FUNCTION_BLOCK "FB_BreakDetector_V1.00"   // FB20, LAD
{ S7_Optimized_Access := 'TRUE' }
VERSION : 0.1
   VAR_INPUT
      IN_xCycleON : Bool;   // Cycle ON
      IN_xCycleONDel : Bool;   // Delayed cycle ON signal
      IN_xGeneralReset : Bool;   // General reset
      IN_xResetAlarms : Bool;   // Reset alarms
      IN_xFaultsEnabled : Bool;   // Faults enabled
      IN_dNumUsedPhoto : DInt;   // Number of used photocell
      IN_dIndexBreakMachine : DInt;   // Index break machine on buffer
      INPUT : Struct   // Digital inputs
         xPowerSupplyControl : Bool;   // Power supply control
         xConnectorONOp : Bool;   // Control connector ON operator side
         xConnectorONOppoOp : Bool;   // Control connector ON opposite operator side
         xButtonAlarmOFF : Bool;   // Reset horn alarm
         rgxPhotoStatus : Array[0..#CONST_DMAXPHOTOCELL_IND] of Bool;   // Photocell status
      END_STRUCT;
   END_VAR
   VAR_OUTPUT
      OUTPUT : Struct
         xLampBreakAlarm : Bool;   // HL.Break alam
         xSirenBreakAlarm : Bool;   // HA.Break alam
      END_STRUCT;
   END_VAR
   VAR_IN_OUT
      INO_tEncoder : "UDT_Encoder";   // Encoder data
      INO_tRibbon : "UDT_RibbonData";   // Ribbona data
      INO_tFBAddDefect : "FB_Defects_Add_V1.00";   // Add defect
      INO_xDefectBufferFull : Bool;   // Defect buffer full
   END_VAR
   VAR RETAIN
      tHMW : Struct   // HMI Write
         dMinBreakSize_cmm : DInt;   // Minimum breaksize [mm/100] {mm/100|mm|0|1000|O}
         rgxEnabledPhotocell : Array[0..#CONST_DMAXPHOTOCELL_IND] of Bool;   // Photocell abilitation (1=Disabled 3=Enabled) {X|X|X|X|O}
         dDistanceSnaproll_cmm : DInt;   // Distance from snaproll [mm/100] {mm/100|mm|0|60000|O}
         xUpdateDistanceSnap : Bool;   // Update distance from snaproll {X|X|X|X|O}
      END_STRUCT;
      tHMR : Struct   // HMI Read
         dStatus : DInt;   // Status (1=Idle 3=Run 5= Glass break 7=Anomaly) {X|X|X|X|O}
         dDistanceSnaproll_cmm : DInt;   // Distance from snaproll [mm/100] {mm/100|mm|0|60000|O}
         rgxPhotoStatus : Array[0..#CONST_DMAXPHOTOCELL_IND] of Bool;   // Photocell status (0=OFF 1=ON) {X|X|X|X|O}
         rgdPhotoAbilitation : Array[0..#CONST_DMAXPHOTOCELL_IND] of DInt;   // Photocell abilitation (1=Disabled 3=Enabled) {X|X|X|X|O}
      END_STRUCT;
   END_VAR
   VAR
      tALM : Struct   // HMI Alarms
         tS : Struct   // Stopping faults machine
            xPowerSupplyControl : Bool;   // Power supply control {X|X|X|X|O}
            xConnectorONOpSide : Bool;   // Connector ON operator side {X|X|X|X|O}
            xConnectorONOppoOpSide : Bool;   // Connector ON opposite operator side {X|X|X|X|O}
            xSpare_3 : Bool;
            xSpare_4 : Bool;
            xSpare_5 : Bool;
            xSpare_6 : Bool;
            xSpare_7 : Bool;
            xSpare_8 : Bool;
            xSpare_9 : Bool;
            xSpare_10 : Bool;
            xSpare_11 : Bool;
            xSpare_12 : Bool;
            xSpare_13 : Bool;
            xSpare_14 : Bool;
            xSpare_15 : Bool;
            xSpare_16 : Bool;
            xSpare_17 : Bool;
            xSpare_18 : Bool;
            xSpare_19 : Bool;
            xSpare_20 : Bool;
            xSpare_21 : Bool;
            xSpare_22 : Bool;
            xSpare_23 : Bool;
            xSpare_24 : Bool;
            xSpare_25 : Bool;
            xSpare_26 : Bool;
            xSpare_27 : Bool;
            xSpare_28 : Bool;
            xSpare_29 : Bool;
            xSpare_30 : Bool;
            xSpare_31 : Bool;
         END_STRUCT;
         tF : Struct   // Faults
            xGlassBreakPhotocell1 : Bool;   // Glass break on photocell #1
            xGlassBreakPhotocell2 : Bool;   // Glass break on photocell #2
            xGlassBreakPhotocell3 : Bool;   // Glass break on photocell #3
            xGlassBreakPhotocell4 : Bool;   // Glass break on photocell #4
            xGlassBreakPhotocell5 : Bool;   // Glass break on photocell #5
            xGlassBreakPhotocell6 : Bool;   // Glass break on photocell #6
            xGlassBreakPhotocell7 : Bool;   // Glass break on photocell #7
            xGlassBreakPhotocell8 : Bool;   // Glass break on photocell #8
            xGlassBreakPhotocell9 : Bool;   // Glass break on photocell #9
            xGlassBreakPhotocell10 : Bool;   // Glass break on photocell #10
            xGlassBreakPhotocell11 : Bool;   // Glass break on photocell #11
            xGlassBreakPhotocell12 : Bool;   // Glass break on photocell #12
            xGlassBreakPhotocell13 : Bool;   // Glass break on photocell #13
            xGlassBreakPhotocell14 : Bool;   // Glass break on photocell #14
            xGlassBreakPhotocell15 : Bool;   // Glass break on photocell #15
            xGlassBreakPhotocell16 : Bool;   // Glass break on photocell #16
            xGlassBreakPhotocell17 : Bool;   // Glass break on photocell #17
            xGlassBreakPhotocell18 : Bool;   // Glass break on photocell #18
            xGlassBreakPhotocell19 : Bool;   // Glass break on photocell #19
            xGlassBreakPhotocell20 : Bool;   // Glass break on photocell #20
            xGlassBreakPhotocell21 : Bool;   // Glass break on photocell #21
            xGlassBreakPhotocell22 : Bool;   // Glass break on photocell #22
            xGlassBreakPhotocell23 : Bool;   // Glass break on photocell #23
            xGlassBreakPhotocell24 : Bool;   // Glass break on photocell #24
            xGlassBreakPhotocell25 : Bool;   // Glass break on photocell #25
            xGlassBreakPhotocell26 : Bool;   // Glass break on photocell #26
            xGlassBreakPhotocell27 : Bool;   // Glass break on photocell #27
            xGlassBreakPhotocell28 : Bool;   // Glass break on photocell #28
            xGlassBreakPhotocell29 : Bool;   // Glass break on photocell #29
            xGlassBreakPhotocell30 : Bool;   // Glass break on photocell #30
            xGlassBreakPhotocell31 : Bool;   // Glass break on photocell #31
            xGlassBreakPhotocell32 : Bool;   // Glass break on photocell #32
         END_STRUCT;
         tW : Struct   // Warnings
            xSpare_0 : Bool;
            xSpare_1 : Bool;
            xSpare_2 : Bool;
            xSpare_3 : Bool;
            xSpare_4 : Bool;
            xSpare_5 : Bool;
            xSpare_6 : Bool;
            xSpare_7 : Bool;
            xSpare_8 : Bool;
            xSpare_9 : Bool;
            xSpare_10 : Bool;
            xSpare_11 : Bool;
            xSpare_12 : Bool;
            xSpare_13 : Bool;
            xSpare_14 : Bool;
            xSpare_15 : Bool;
            xSpare_16 : Bool;
            xSpare_17 : Bool;
            xSpare_18 : Bool;
            xSpare_19 : Bool;
            xSpare_20 : Bool;
            xSpare_21 : Bool;
            xSpare_22 : Bool;
            xSpare_23 : Bool;
            xSpare_24 : Bool;
            xSpare_25 : Bool;
            xSpare_26 : Bool;
            xSpare_27 : Bool;
            xSpare_28 : Bool;
            xSpare_29 : Bool;
            xSpare_30 : Bool;
            xSpare_31 : Bool;
         END_STRUCT;
      END_STRUCT;
      ST_xOutputEnable : Bool;   // Output enable
      ST_xStoppedFaults : Bool;   // Stopped faults
      ST_xFaults : Bool;   // Faults
      ST_xWarning : Bool;   // Warnings
      AUX_rgxLastPhotoState : Array[0..#CONST_DMAXPHOTOCELL_IND] of Bool;   // Last photocell status
      AUX_xGlassBreak : Bool;   // Glass break in progress
      AUX_xGlassBreakInGoing : Bool;   // Glass break ingoing
      AUX_dCounterOnBreak_cmm : DInt;   // Encoder counter on glass break front
      AUX_dLastInsertDefectPos_cmm : DInt;   // Last inserted defect position [mm/100]
      OSR_xGlassBreak : Bool;   // OSR glasss break
   END_VAR
   VAR_TEMP
      TMP_dwValue : DWord;
      TMP_dIndex : DInt;
      TMP_dNumUsedPhotocell : DInt;
      TMP_xGlassBreak : Bool;
      TMP_xAtLeastOnePhoto : Bool;
      TMP_dEncDef_cmm : DInt;
   END_VAR
   VAR CONSTANT
      CONST_DMAXPHOTOCELL : DInt := 32;   // Maximum number of photocell
      CONST_DMAXPHOTOCELL_IND : DInt := 31;   // Maximum number of photocell index (Always -1)
      CONST_DGLASSBREAK_CLASS : DInt := 21;   // Glass break used class
      CONST_DGLASSBREAK_SUBTYPE : DInt := 1002;   // Glass break subtype
      CONST_DGLASSBREAK_DEFECT_WIDTH_CMM : DInt := 366000;   // Defect width [mm/100]
      CONST_DGLASSBREAK_DEFECT_GAP_CMM : DInt := 40000;   // Glass break defect gap [mm/100]
      CONST_DGLASSBREAK_LASTDEFECT_LENGTH_CMM : DInt := 50000;   // Last defect on glass break length [mm/100]
   END_VAR
   VAR_TEMP   // added for the SCL form of the ladder/FBD networks
      _w1 : Bool;
   END_VAR
BEGIN

REGION Network 1: ####_CONSTANTS_####
END_REGION

REGION Network 2: ####_MATCH_####
END_REGION

REGION Network 3 (SCL): ### SIMULATION ###
   IF "SIMULATION_ACTIVE" THEN
       #INPUT.xConnectorONOp := TRUE;
       #INPUT.xConnectorONOppoOp := TRUE;
       #INPUT.xPowerSupplyControl := TRUE;
    //   #INPUT.rgxPhotoStatus[0] := 1;
   //    #INPUT.rgxPhotoStatus[1] := 1;
   //    #INPUT.rgxPhotoStatus[2] := 1;
   //    #INPUT.rgxPhotoStatus[3] := 1;
    //   #INPUT.rgxPhotoStatus[4] := 1;
     //  #INPUT.rgxPhotoStatus[5] := 1;
    //   #INPUT.rgxPhotoStatus[6] := 1;
     //  #INPUT.rgxPhotoStatus[7] := 1;
     //  #INPUT.rgxPhotoStatus[8] := 1;
      // #INPUT.rgxPhotoStatus[9] := 1;
   END_IF;
END_REGION

REGION Network 4 (SCL): Evaluate number of used photocell
   #TMP_dNumUsedPhotocell := #IN_dNumUsedPhoto;

   IF #TMP_dNumUsedPhotocell > #CONST_DMAXPHOTOCELL THEN
       #TMP_dNumUsedPhotocell := #CONST_DMAXPHOTOCELL;
   ELSIF #TMP_dNumUsedPhotocell < 0 THEN
       #TMP_dNumUsedPhotocell := 0;
   END_IF;
END_REGION

REGION Network 5 (SCL): Reset all the pending status
   IF #IN_xGeneralReset THEN
       #AUX_xGlassBreak := FALSE;
       #AUX_xGlassBreakInGoing := FALSE;
       #AUX_dCounterOnBreak_cmm := 0;

       FOR #TMP_dIndex := 0 TO #TMP_dNumUsedPhotocell - 1 DO
           #AUX_rgxLastPhotoState[#TMP_dIndex] := FALSE;
       END_FOR;

   END_IF;
END_REGION

REGION Network 6: ####_HMI_LOGICS_####
END_REGION

REGION Network 7 (SCL): Manage HMI Logics
   FOR #TMP_dIndex := 0 TO #TMP_dNumUsedPhotocell - 1 DO

       (*  IF #tHMW.rgxEnabledPhotocell[#TMP_dIndex] THEN
           #tHMW.rgxEnabledPhotocell[#TMP_dIndex] := FALSE;
           #tHMR.rgdPhotoAbilitation[#TMP_dIndex] := 3;
       END_IF;

       IF #tHMW.rgxDisablePhotocell[#TMP_dIndex] THEN
           #tHMW.rgxDisablePhotocell[#TMP_dIndex] := FALSE;
           #tHMR.rgdPhotoAbilitation[#TMP_dIndex] := 1;
       END_IF; 
       IF #tHMW.rgxEnabledPhotocell[#TMP_dIndex] THEN
           #tHMW.rgxEnabledPhotocell[#TMP_dIndex] := FALSE;
           #tHMR.rgdPhotoAbilitation[#TMP_dIndex] := 3;
       END_IF;*)

       IF #tHMW.rgxEnabledPhotocell[#TMP_dIndex] =1 THEN

           #tHMR.rgdPhotoAbilitation[#TMP_dIndex] := 3;
       ELSE
           #tHMR.rgdPhotoAbilitation[#TMP_dIndex] := 1;
       END_IF;


   END_FOR;

   IF #tHMW.xUpdateDistanceSnap  THEN

       #tHMW.xUpdateDistanceSnap := FALSE;
       #tHMR.dDistanceSnaproll_cmm := #tHMW.dDistanceSnaproll_cmm;
       #INO_tRibbon.rgtGlassBreak[#IN_dIndexBreakMachine].dDistSnapRoll_cmm := #tHMR.dDistanceSnaproll_cmm;

   END_IF;
END_REGION

REGION Network 8: ####_ALARMS_####
END_REGION

REGION Network 9 (SCL): Reset alarms
   IF #IN_xResetAlarms THEN

       #TMP_dwValue := 0;

       SCATTER(IN:=#TMP_dwValue,
               OUT=>#tALM.tS);

       SCATTER(IN:=#TMP_dwValue,
               OUT=>#tALM.tF);

       SCATTER(IN:=#TMP_dwValue,
               OUT=>#tALM.tW);


   END_IF;
END_REGION

REGION Network 10: Power supply control
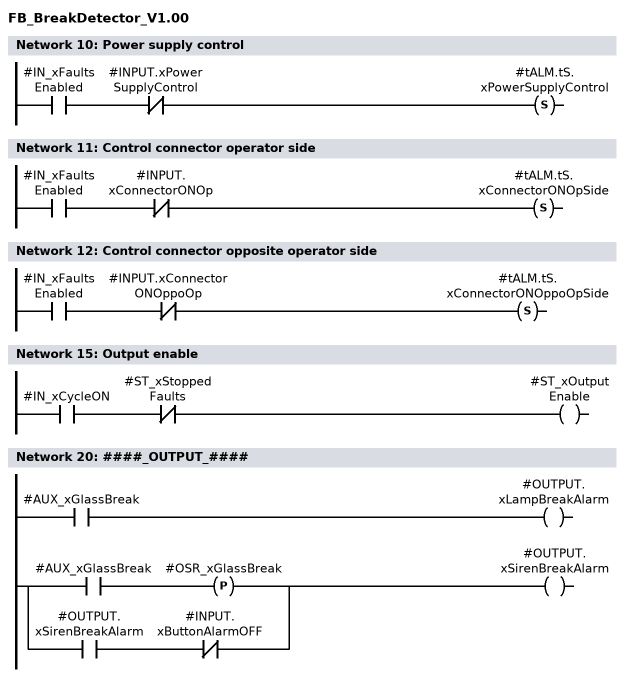
   RUNG wire#powerrail
      Contact( #IN_xFaultsEnabled )
      I_Contact( #INPUT.xPowerSupplyControl )
      S_Coil( #tALM.tS.xPowerSupplyControl )
   END_RUNG
   // the same network as SCL:
   IF #IN_xFaultsEnabled AND NOT #INPUT.xPowerSupplyControl THEN
       #tALM.tS.xPowerSupplyControl := TRUE;
   END_IF;
END_REGION

REGION Network 11: Control connector operator side
   RUNG wire#powerrail
      Contact( #IN_xFaultsEnabled )
      I_Contact( #INPUT.xConnectorONOp )
      S_Coil( #tALM.tS.xConnectorONOpSide )
   END_RUNG
   // the same network as SCL:
   IF #IN_xFaultsEnabled AND NOT #INPUT.xConnectorONOp THEN #tALM.tS.xConnectorONOpSide := TRUE; END_IF;
END_REGION

REGION Network 12: Control connector opposite operator side
   RUNG wire#powerrail
      Contact( #IN_xFaultsEnabled )
      I_Contact( #INPUT.xConnectorONOppoOp )
      S_Coil( #tALM.tS.xConnectorONOppoOpSide )
   END_RUNG
   // the same network as SCL:
   IF #IN_xFaultsEnabled AND NOT #INPUT.xConnectorONOppoOp THEN
       #tALM.tS.xConnectorONOppoOpSide := TRUE;
   END_IF;
END_REGION

REGION Network 13 (SCL): Calculate comulative statuses
       GATHER(IN:=#tALM.tS,
              OUT=>#TMP_dwValue);

       IF #TMP_dwValue <> 0 THEN
           #ST_xStoppedFaults := TRUE;
       ELSE
           #ST_xStoppedFaults := FALSE;
       END_IF;

       GATHER(IN:=#tALM.tF,
              OUT=>#TMP_dwValue);

       IF #TMP_dwValue <> 0 THEN
           #ST_xFaults := TRUE;
       ELSE
           #ST_xFaults := FALSE;
       END_IF;

       GATHER(IN:=#tALM.tW,
              OUT=>#TMP_dwValue);

       IF #TMP_dwValue <> 0 THEN
           #ST_xWarning := TRUE;
       ELSE
           #ST_xWarning := FALSE;
       END_IF;
END_REGION

REGION Network 14: ####_STATUSES_####
END_REGION

REGION Network 15: Output enable
   RUNG wire#powerrail
      Contact( #IN_xCycleON )
      I_Contact( #ST_xStoppedFaults )
      Coil( #ST_xOutputEnable )
   END_RUNG
   // the same network as SCL:
   #ST_xOutputEnable := #IN_xCycleON AND NOT #ST_xStoppedFaults;
END_REGION

REGION Network 16: ### PHASES AND LOGICS ###
END_REGION

REGION Network 17 (SCL): Evaluate glass break
   #TMP_xGlassBreak := FALSE;

   FOR #TMP_dIndex := 0 TO #TMP_dNumUsedPhotocell - 1 DO

       IF #INPUT.rgxPhotoStatus[#TMP_dIndex] = FALSE AND #tHMR.rgdPhotoAbilitation[#TMP_dIndex] = 3 AND #ST_xOutputEnable THEN
           #TMP_xGlassBreak := TRUE;
       END_IF;    

       #AUX_rgxLastPhotoState[#TMP_dIndex] := #INPUT.rgxPhotoStatus[#TMP_dIndex];

   END_FOR;

   //In case of glassbreak front up, evaluate the space elapse from the other front
   IF (#TMP_xGlassBreak = TRUE) AND (#AUX_xGlassBreak = FALSE) AND (#AUX_xGlassBreakInGoing = FALSE) THEN
       #AUX_dCounterOnBreak_cmm := #INO_tEncoder.dActualEncoderCounter_cmm;
       #AUX_xGlassBreakInGoing := TRUE;
   ELSIF (#TMP_xGlassBreak = FALSE) THEN
       #AUX_xGlassBreakInGoing := FALSE;

       //If glass break was true, update the front off
       IF (#AUX_xGlassBreak = TRUE) THEN

           #INO_tRibbon.rgtGlassBreakUpdate[#IN_dIndexBreakMachine].tData.dEncoderValue_cmm := 0;
           #INO_tRibbon.rgtGlassBreakUpdate[#IN_dIndexBreakMachine].tData.xGlassBreak := FALSE;

           #TMP_dwValue := 0;
           SCATTER(IN:=#TMP_dwValue, OUT=>#INO_tRibbon.rgtGlassBreakUpdate[#IN_dIndexBreakMachine].tData.rgxBreakMask);

           #INO_tRibbon.rgtGlassBreakUpdate[#IN_dIndexBreakMachine].tData.xUpdateDataBPSA := TRUE;
           #INO_tRibbon.rgtGlassBreakUpdate[#IN_dIndexBreakMachine].tData.xUpdateDataBPSB := TRUE;
           #INO_tRibbon.rgtGlassBreakUpdate[#IN_dIndexBreakMachine].xUpdateRequest := TRUE;

           //Insert defect on the buffer to close the glass break
           #INO_tFBAddDefect(IN_dClass:=#CONST_DGLASSBREAK_CLASS,
                         IN_dSubType:=#CONST_DGLASSBREAK_SUBTYPE,
                         IN_dXPosition_cmm:=#INO_tEncoder.dActualEncoderCounter_cmm + #tHMR.dDistanceSnaproll_cmm,
                         IN_dYPosition_cmm:= #CONST_DGLASSBREAK_DEFECT_WIDTH_CMM / -2,
                         IN_dTotalLength_um:= #CONST_DGLASSBREAK_LASTDEFECT_LENGTH_CMM * 10,
                         IN_dTotalWidth_um:=#CONST_DGLASSBREAK_DEFECT_WIDTH_CMM * 10,
                         IN_dCoreLength_um := #CONST_DGLASSBREAK_LASTDEFECT_LENGTH_CMM * 10,
                         IN_dCoreWidth_um:=#CONST_DGLASSBREAK_DEFECT_WIDTH_CMM * 10,
                         IN_dDistLength_um := #CONST_DGLASSBREAK_LASTDEFECT_LENGTH_CMM * 10,
                         IN_dDistWidth_um:=#CONST_DGLASSBREAK_DEFECT_WIDTH_CMM * 10,
                         IN_dOptValue_mdptr:=0,
                         OUT_xBufferFull => #INO_xDefectBufferFull,
                         IN_strDefectID:='GLASS_BREAK');

       END_IF;

       #AUX_xGlassBreak := FALSE;

   END_IF;

   //If glass break ingoing evaluate the space, if space greather than filter activate the break
   IF (#AUX_xGlassBreakInGoing = TRUE) AND 
           (#INO_tEncoder.dActualEncoderCounter_cmm - #AUX_dCounterOnBreak_cmm) >= #tHMW.dMinBreakSize_cmm THEN

       #AUX_xGlassBreakInGoing := FALSE;
       #AUX_xGlassBreak := TRUE;

       //Insert the break on the buffer
       #INO_tRibbon.rgtGlassBreakUpdate[#IN_dIndexBreakMachine].tData.dEncoderValue_cmm := 0;
       #INO_tRibbon.rgtGlassBreakUpdate[#IN_dIndexBreakMachine].tData.xGlassBreak := TRUE;

       #TMP_dwValue := 0;

       SCATTER(IN:=#TMP_dwValue, OUT=>#INO_tRibbon.rgtGlassBreakUpdate[#IN_dIndexBreakMachine].tData.rgxBreakMask);

       FOR #TMP_dIndex := 0 TO #TMP_dNumUsedPhotocell - 1 DO
           IF #INPUT.rgxPhotoStatus[#TMP_dIndex] = FALSE AND #tHMR.rgdPhotoAbilitation[#TMP_dIndex] = 3 THEN
               #INO_tRibbon.rgtGlassBreakUpdate[#IN_dIndexBreakMachine].tData.rgxBreakMask[#TMP_dIndex] := TRUE;
           ELSE                
               #INO_tRibbon.rgtGlassBreakUpdate[#IN_dIndexBreakMachine].tData.rgxBreakMask[#TMP_dIndex] := FALSE;
           END_IF;
       END_FOR;

       #INO_tRibbon.rgtGlassBreakUpdate[#IN_dIndexBreakMachine].tData.xUpdateDataBPSA := TRUE;
       #INO_tRibbon.rgtGlassBreakUpdate[#IN_dIndexBreakMachine].tData.xUpdateDataBPSB := TRUE;

       #INO_tRibbon.rgtGlassBreakUpdate[#IN_dIndexBreakMachine].xUpdateRequest := TRUE;

       //Insert defect on the buffer
       #INO_tFBAddDefect(IN_dClass:=#CONST_DGLASSBREAK_CLASS,
                         IN_dSubType:=#CONST_DGLASSBREAK_SUBTYPE,
                         IN_dXPosition_cmm:=#AUX_dCounterOnBreak_cmm  + #tHMR.dDistanceSnaproll_cmm,
                         IN_dYPosition_cmm:= #CONST_DGLASSBREAK_DEFECT_WIDTH_CMM / -2,
                         IN_dTotalLength_um:= 1000,
                         IN_dTotalWidth_um:=#CONST_DGLASSBREAK_DEFECT_WIDTH_CMM * 10,
                         IN_dCoreLength_um := 1000,
                         IN_dCoreWidth_um:=#CONST_DGLASSBREAK_DEFECT_WIDTH_CMM * 10,
                         IN_dDistLength_um := 1000,
                         IN_dDistWidth_um:=#CONST_DGLASSBREAK_DEFECT_WIDTH_CMM * 10,
                         IN_dOptValue_mdptr:=0,
                         OUT_xBufferFull => #INO_xDefectBufferFull,
                         IN_strDefectID:='GLASS_BREAK');

       #AUX_dLastInsertDefectPos_cmm := #AUX_dCounterOnBreak_cmm  + #tHMR.dDistanceSnaproll_cmm;

   END_IF;
END_REGION

REGION Network 18 (SCL): Insert defect in according the glass break
   IF (#AUX_xGlassBreak) THEN

       #TMP_dEncDef_cmm := #INO_tEncoder.dActualEncoderCounter_cmm + #tHMR.dDistanceSnaproll_cmm;

       IF (#TMP_dEncDef_cmm - #AUX_dLastInsertDefectPos_cmm) > #CONST_DGLASSBREAK_DEFECT_GAP_CMM THEN

       #AUX_dLastInsertDefectPos_cmm := #INO_tEncoder.dActualEncoderCounter_cmm + #tHMR.dDistanceSnaproll_cmm;    
       //Insert defect on the buffer
       #INO_tFBAddDefect(IN_dClass:= #CONST_DGLASSBREAK_CLASS,
                         IN_dSubType:= #CONST_DGLASSBREAK_SUBTYPE,
                         IN_dXPosition_cmm:= #AUX_dLastInsertDefectPos_cmm,
                         IN_dYPosition_cmm:= #CONST_DGLASSBREAK_DEFECT_WIDTH_CMM / -2,
                         IN_dTotalLength_um:= 1000,
                         IN_dTotalWidth_um:= #CONST_DGLASSBREAK_DEFECT_WIDTH_CMM * 10,
                         IN_dCoreLength_um := 1000,
                         IN_dCoreWidth_um:=#CONST_DGLASSBREAK_DEFECT_WIDTH_CMM * 10,
                         IN_dDistLength_um := 1000,
                         IN_dDistWidth_um:=#CONST_DGLASSBREAK_DEFECT_WIDTH_CMM * 10,
                         IN_dOptValue_mdptr:=0,
                         OUT_xBufferFull => #INO_xDefectBufferFull,
                         IN_strDefectID:='GLASS_BREAK');

       END_IF;

   END_IF;
END_REGION

REGION Network 19 (SCL): ### HMI STATUS ###
   //At least one photocell enabled
   #TMP_xAtLeastOnePhoto := FALSE;
   FOR #TMP_dIndex := 0 TO #TMP_dNumUsedPhotocell - 1 DO

       IF #tHMR.rgdPhotoAbilitation[#TMP_dIndex] = 3 THEN 
           #TMP_xAtLeastOnePhoto := TRUE;
           EXIT;    
       END_IF;

   END_FOR;

   FOR #TMP_dIndex := 0 TO #TMP_dNumUsedPhotocell - 1 DO

       #tHMR.rgxPhotoStatus[#TMP_dIndex] := #INPUT.rgxPhotoStatus[#TMP_dIndex];

   END_FOR;

   //Calculate status
   IF #ST_xStoppedFaults THEN
       #tHMR.dStatus := 7;
   ELSIF #AUX_xGlassBreak THEN
       #tHMR.dStatus := 5;
   ELSIF #TMP_xAtLeastOnePhoto THEN
       #tHMR.dStatus := 3;
   ELSE
       #tHMR.dStatus := 1;
   END_IF;
END_REGION

REGION Network 20: ####_OUTPUT_####
   RUNG wire#powerrail
      Contact( #AUX_xGlassBreak )
      Coil( #OUTPUT.xLampBreakAlarm )
   END_RUNG
   RUNG wire#powerrail
      Contact( #AUX_xGlassBreak )
      P_Trig( #OSR_xGlassBreak )
      wire#w1
      Coil( #OUTPUT.xSirenBreakAlarm )
   END_RUNG
   RUNG wire#powerrail
      Contact( #OUTPUT.xSirenBreakAlarm )
      I_Contact( #INPUT.xButtonAlarmOFF )
   END_RUNG wire#w1
   // the same network as SCL:
   #OUTPUT.xLampBreakAlarm := #AUX_xGlassBreak;
   #_w1 := #AUX_xGlassBreak AND NOT #OSR_xGlassBreak;   // rising edge
   #OSR_xGlassBreak := #AUX_xGlassBreak;
   #OUTPUT.xSirenBreakAlarm := #_w1 OR (#OUTPUT.xSirenBreakAlarm AND NOT #INPUT.xButtonAlarmOFF);
END_REGION
END_FUNCTION_BLOCK

// folder: 03_Programs_Logics/MCC1201/19_Breaker

FUNCTION_BLOCK "FB_BreakerM206_V1.00"   // FB29, LAD
{ S7_Optimized_Access := 'TRUE' }
VERSION : 0.1
   VAR_INPUT
      IN_xCycleON : Bool;   // Cycle ON
      IN_xCycleONDel : Bool;   // Delayed cycle ON signal
      IN_xGeneralReset : Bool;   // General reset
      IN_xResetAlarms : Bool;   // Reset alarms
      IN_xFaultsEnabled : Bool;   // Faults enabled
      IN_xDropConveyorDown : Bool;   // Run request - drop conveyor down
      INPUT : Struct   // Digital inputs
         xConditionOKFromCulletSystem : Bool;   // X.Condition ok cullet system
         xBreakerRotationControl : Bool;   // SQ.Braker rotation feedback
         xProtectionBreakerRotation : Bool;   // Q.Protection breaker rotation
         xFeedbackRotationKM : Bool;
      END_STRUCT;
   END_VAR
   VAR_OUTPUT
      OUTPUT : Struct
         xBreakerRun : Bool;   // Breaker start
         xToScrapingUnderZ200 : Bool;
         xHlScrapinglineReady : Bool;
         xHlScrapinglineNotReady : Bool;
      END_STRUCT;
   END_VAR
   VAR_IN_OUT
      INO_tOBInitialize : "GP_OB_Initialize";   // OB Initialize
   END_VAR
   VAR
      tHMW : Struct   // HMI Write
         tManCmd : Struct
            xRun : Bool := false;   // Manual run {x|x|x|x|O}
         END_STRUCT;
         xEnableManualCommand : Bool;   // Enable Manual command {x|x|x|x|O}
         xEnableRunAlwaysModeBreaker : Bool;   // Enable run always breaker {x|x|x|x|O}
         dBreakerRetainTime_s : DInt;   // Breaker retain command after rise {ms|s|0|120|O}
      END_STRUCT;
      tHMR : Struct   // HMI Read
         tManCmd : Struct
            xRunFdbk : Bool;   // Manual run fdbk {x|x|x|x|O}
         END_STRUCT;
         xManualCommandEnabled : Bool;   // Manual Command enabled {x|x|x|x|O}
         xEnabledRunAlwaysModeBreaker : Bool;   // Enabled run always breaker {x|x|x|x|O}
         dStatus : DInt;   // Status (1=Idle 3=Run 7=Anomaly) {X|X|X|X|O}
      END_STRUCT;
      tALM : Struct   // HMI Alarms
         tS : Struct   // Stopping faults machine
            xSpare_1 : Bool;
            xConditionOKCulletSystem : Bool;   // Condition OK from cullet system {X|X|X|X|O}
            xBreakerRotationFeedback : Bool;   // A406SQ1.Breaker rotation feedback {X|X|X|X|O}
            xBreakerKmRotationFeedback : Bool;
            xSpare_3 : Bool;
            xProtectionBreakerRotation : Bool;   // QM.Protection breaker rotation {X|X|X|X|O}
            xSpare_4 : Bool;
            xSpare_5 : Bool;
            xSpare_6 : Bool;
            xSpare_7 : Bool;
            xSpare_8 : Bool;
            xSpare_9 : Bool;
            xSpare_10 : Bool;
            xSpare_11 : Bool;
            xSpare_14 : Bool;
            xSpare_15 : Bool;
            xSpare_16 : Bool;
            xSpare_17 : Bool;
            xSpare_18 : Bool;
            xSpare_19 : Bool;
            xSpare_20 : Bool;
            xSpare_21 : Bool;
            xSpare_22 : Bool;
            xSpare_23 : Bool;
            xSpare_24 : Bool;
            xSpare_25 : Bool;
            xSpare_26 : Bool;
            xSpare_27 : Bool;
            xSpare_28 : Bool;
            xSpare_29 : Bool;
            xSpare_30 : Bool;
            xSpare_31 : Bool;
         END_STRUCT;
         tF : Struct   // Faults
            xSpare_0 : Bool;
            xSpare_1 : Bool;
            xSpare_2 : Bool;
            xSpare_3 : Bool;
            xSpare_4 : Bool;
            xSpare_5 : Bool;
            xSpare_6 : Bool;
            xSpare_7 : Bool;
            xSpare_8 : Bool;
            xSpare_9 : Bool;
            xSpare_10 : Bool;
            xSpare_11 : Bool;
            xSpare_12 : Bool;
            xSpare_13 : Bool;
            xSpare_14 : Bool;
            xSpare_15 : Bool;
            xSpare_16 : Bool;
            xSpare_17 : Bool;
            xSpare_18 : Bool;
            xSpare_19 : Bool;
            xSpare_20 : Bool;
            xSpare_21 : Bool;
            xSpare_22 : Bool;
            xSpare_23 : Bool;
            xSpare_24 : Bool;
            xSpare_25 : Bool;
            xSpare_26 : Bool;
            xSpare_27 : Bool;
            xSpare_28 : Bool;
            xSpare_29 : Bool;
            xSpare_30 : Bool;
            xSpare_31 : Bool;
         END_STRUCT;
         tW : Struct   // Warnings
            xSpare_0 : Bool;
            xSpare_1 : Bool;
            xSpare_2 : Bool;
            xSpare_3 : Bool;
            xSpare_4 : Bool;
            xSpare_5 : Bool;
            xSpare_6 : Bool;
            xSpare_7 : Bool;
            xSpare_8 : Bool;
            xSpare_9 : Bool;
            xSpare_10 : Bool;
            xSpare_11 : Bool;
            xSpare_12 : Bool;
            xSpare_13 : Bool;
            xSpare_14 : Bool;
            xSpare_15 : Bool;
            xSpare_16 : Bool;
            xSpare_17 : Bool;
            xSpare_18 : Bool;
            xSpare_19 : Bool;
            xSpare_20 : Bool;
            xSpare_21 : Bool;
            xSpare_22 : Bool;
            xSpare_23 : Bool;
            xSpare_24 : Bool;
            xSpare_25 : Bool;
            xSpare_26 : Bool;
            xSpare_27 : Bool;
            xSpare_28 : Bool;
            xSpare_29 : Bool;
            xSpare_30 : Bool;
            xSpare_31 : Bool;
         END_STRUCT;
      END_STRUCT;
      ST_xManualMode : Bool;   // Manual mode
      ST_xOutputEnable : Bool;   // Output enable
      ST_xCondOkMan : Bool;   // Condition ok manual command
      ST_xStoppedFaults : Bool;   // Stopped faults
      ST_xFaults : Bool;   // Faults
      ST_xWarning : Bool;   // Warnings
      AUX_tmOFF_RunRetain : "UDT_IECTOFF_V1.00";   // Feedback retain
      AUX_tmON_FeedbackRotAno : "UDT_IECTON_V1.00";   // Feedback rotation anomaly
      AUX_tmON_FeedbackKMRotAno : "UDT_IECTON_V1.00";   // Feedback rotation anomaly
   END_VAR
   VAR_TEMP
      TMP_dwValue : DWord;
   END_VAR
   VAR CONSTANT
      CONST_DSTATUS_ANOMALY : DInt := 7;
      CONST_DSTATUS_RUN : DInt := 3;
      CONST_DSTATUS_IDLE : DInt := 1;
   END_VAR
   VAR_TEMP   // added for the SCL form of the ladder/FBD networks
      _w1 : Bool;
   END_VAR
BEGIN

REGION Network 1: ####_CONSTANTS_####
END_REGION

REGION Network 2 (SCL): ### SIMULATION ###
   IF "SIMULATION_ACTIVE" THEN

       #INPUT.xConditionOKFromCulletSystem := TRUE;
       #INPUT.xBreakerRotationControl := #OUTPUT.xBreakerRun;
       #INPUT.xProtectionBreakerRotation := TRUE;

   END_IF;
END_REGION

REGION Network 3: ####_MATCH_####
END_REGION

REGION Network 4: ####_HMI_LOGICS_####
END_REGION

REGION Network 5: Enabled run always breaker
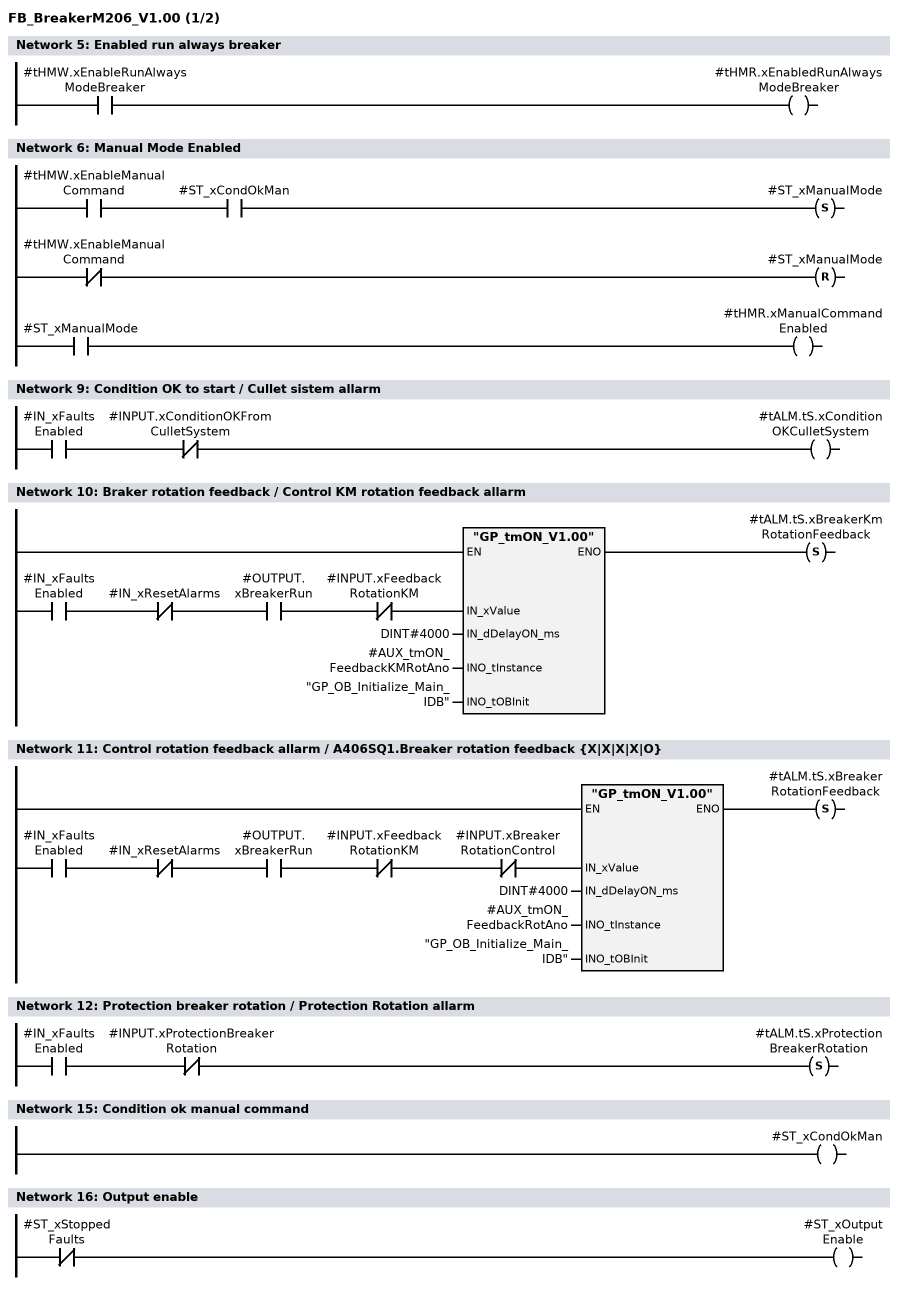
   RUNG wire#powerrail
      Contact( #tHMW.xEnableRunAlwaysModeBreaker )
      Coil( #tHMR.xEnabledRunAlwaysModeBreaker )
   END_RUNG
   // the same network as SCL:
   #tHMR.xEnabledRunAlwaysModeBreaker := #tHMW.xEnableRunAlwaysModeBreaker;
END_REGION

REGION Network 6: Manual Mode Enabled
   RUNG wire#powerrail
      Contact( #tHMW.xEnableManualCommand )
      Contact( #ST_xCondOkMan )
      S_Coil( #ST_xManualMode )
   END_RUNG
   RUNG wire#powerrail
      I_Contact( #tHMW.xEnableManualCommand )
      R_Coil( #ST_xManualMode )
   END_RUNG
   RUNG wire#powerrail
      Contact( #ST_xManualMode )
      Coil( #tHMR.xManualCommandEnabled )
   END_RUNG
   // the same network as SCL:
   IF #tHMW.xEnableManualCommand AND #ST_xCondOkMan THEN #ST_xManualMode := TRUE; END_IF;
   IF NOT #tHMW.xEnableManualCommand THEN #ST_xManualMode := FALSE; END_IF;
   #tHMR.xManualCommandEnabled := #ST_xManualMode;
END_REGION

REGION Network 7: ####_ALARMS_####
END_REGION

REGION Network 8 (SCL): Reset alarms
   IF #IN_xResetAlarms THEN

       #TMP_dwValue := 0;

       SCATTER(IN:=#TMP_dwValue,
               OUT=>#tALM.tS);

       SCATTER(IN:=#TMP_dwValue,
               OUT=>#tALM.tF);

       SCATTER(IN:=#TMP_dwValue,
               OUT=>#tALM.tW);


   END_IF;
END_REGION

REGION Network 9: Condition OK to start / Cullet sistem allarm
   RUNG wire#powerrail
      Contact( #IN_xFaultsEnabled )
      I_Contact( #INPUT.xConditionOKFromCulletSystem )
      Coil( #tALM.tS.xConditionOKCulletSystem )
   END_RUNG
   // the same network as SCL:
   #tALM.tS.xConditionOKCulletSystem := #IN_xFaultsEnabled AND NOT #INPUT.xConditionOKFromCulletSystem;
END_REGION

REGION Network 10: Braker rotation feedback / Control KM rotation feedback allarm
   RUNG wire#powerrail
      "GP_tmON_V1.00"(IN_xValue := wire#w1, IN_dDelayON_ms := DINT#4000, INO_tInstance := #AUX_tmON_FeedbackKMRotAno, INO_tOBInit := "GP_OB_Initialize_Main_IDB")
      S_Coil( #tALM.tS.xBreakerKmRotationFeedback )
   END_RUNG
   RUNG wire#powerrail
      Contact( #IN_xFaultsEnabled )
      I_Contact( #IN_xResetAlarms )
      Contact( #OUTPUT.xBreakerRun )
      I_Contact( #INPUT.xFeedbackRotationKM )
   END_RUNG wire#w1
   // the same network as SCL:
   "GP_tmON_V1.00"(IN_xValue := #IN_xFaultsEnabled AND NOT #IN_xResetAlarms AND #OUTPUT.xBreakerRun AND NOT #INPUT.xFeedbackRotationKM,
                   IN_dDelayON_ms := DINT#4000,
                   INO_tInstance := #AUX_tmON_FeedbackKMRotAno,
                   INO_tOBInit := "GP_OB_Initialize_Main_IDB",
                   ENO => #_w1);
   IF #_w1 THEN #tALM.tS.xBreakerKmRotationFeedback := TRUE; END_IF;
END_REGION

REGION Network 11: Control rotation feedback allarm / A406SQ1.Breaker rotation feedback {X|X|X|X|O}
   RUNG wire#powerrail
      "GP_tmON_V1.00"(IN_xValue := wire#w1, IN_dDelayON_ms := DINT#4000, INO_tInstance := #AUX_tmON_FeedbackRotAno, INO_tOBInit := "GP_OB_Initialize_Main_IDB")
      S_Coil( #tALM.tS.xBreakerRotationFeedback )
   END_RUNG
   RUNG wire#powerrail
      Contact( #IN_xFaultsEnabled )
      I_Contact( #IN_xResetAlarms )
      Contact( #OUTPUT.xBreakerRun )
      I_Contact( #INPUT.xFeedbackRotationKM )
      I_Contact( #INPUT.xBreakerRotationControl )
   END_RUNG wire#w1
   // the same network as SCL:
   "GP_tmON_V1.00"(IN_xValue := #IN_xFaultsEnabled AND NOT #IN_xResetAlarms AND #OUTPUT.xBreakerRun AND NOT #INPUT.xFeedbackRotationKM AND NOT #INPUT.xBreakerRotationControl,
                   IN_dDelayON_ms := DINT#4000,
                   INO_tInstance := #AUX_tmON_FeedbackRotAno,
                   INO_tOBInit := "GP_OB_Initialize_Main_IDB",
                   ENO => #_w1);
   IF #_w1 THEN #tALM.tS.xBreakerRotationFeedback := TRUE; END_IF;
END_REGION

REGION Network 12: Protection breaker rotation / Protection Rotation allarm
   RUNG wire#powerrail
      Contact( #IN_xFaultsEnabled )
      I_Contact( #INPUT.xProtectionBreakerRotation )
      S_Coil( #tALM.tS.xProtectionBreakerRotation )
   END_RUNG
   // the same network as SCL:
   IF #IN_xFaultsEnabled AND NOT #INPUT.xProtectionBreakerRotation THEN
       #tALM.tS.xProtectionBreakerRotation := TRUE;
   END_IF;
END_REGION

REGION Network 13 (SCL): Calculate comulative statuses
       GATHER(IN:=#tALM.tS,
              OUT=>#TMP_dwValue);

       IF #TMP_dwValue <> 0 THEN
           #ST_xStoppedFaults := TRUE;
       ELSE
           #ST_xStoppedFaults := FALSE;
       END_IF;

       GATHER(IN:=#tALM.tF,
              OUT=>#TMP_dwValue);

       IF #TMP_dwValue <> 0 THEN
           #ST_xFaults := TRUE;
       ELSE
           #ST_xFaults := FALSE;
       END_IF;

       GATHER(IN:=#tALM.tW,
              OUT=>#TMP_dwValue);

       IF #TMP_dwValue <> 0 THEN
           #ST_xWarning := TRUE;
       ELSE
           #ST_xWarning := FALSE;
       END_IF;
END_REGION

REGION Network 14: ####_STATUSES_####
END_REGION

REGION Network 15: Condition ok manual command
   RUNG wire#powerrail
      Coil( #ST_xCondOkMan )
   END_RUNG
   // the same network as SCL:
   #ST_xCondOkMan := TRUE;
END_REGION

REGION Network 16: Output enable
   RUNG wire#powerrail
      I_Contact( #ST_xStoppedFaults )
      Coil( #ST_xOutputEnable )
   END_RUNG
   // the same network as SCL:
   #ST_xOutputEnable := NOT #ST_xStoppedFaults;
END_REGION

REGION Network 17 (SCL): ### HMI STATUS ###
   IF #ST_xStoppedFaults THEN
       #tHMR.dStatus := #CONST_DSTATUS_ANOMALY;
   ELSIF #INPUT.xBreakerRotationControl THEN
       #tHMR.dStatus := #CONST_DSTATUS_RUN;
   ELSE
       #tHMR.dStatus := #CONST_DSTATUS_IDLE;
   END_IF;
END_REGION

REGION Network 18: Manual run fdbk {x|x|x|x|O}
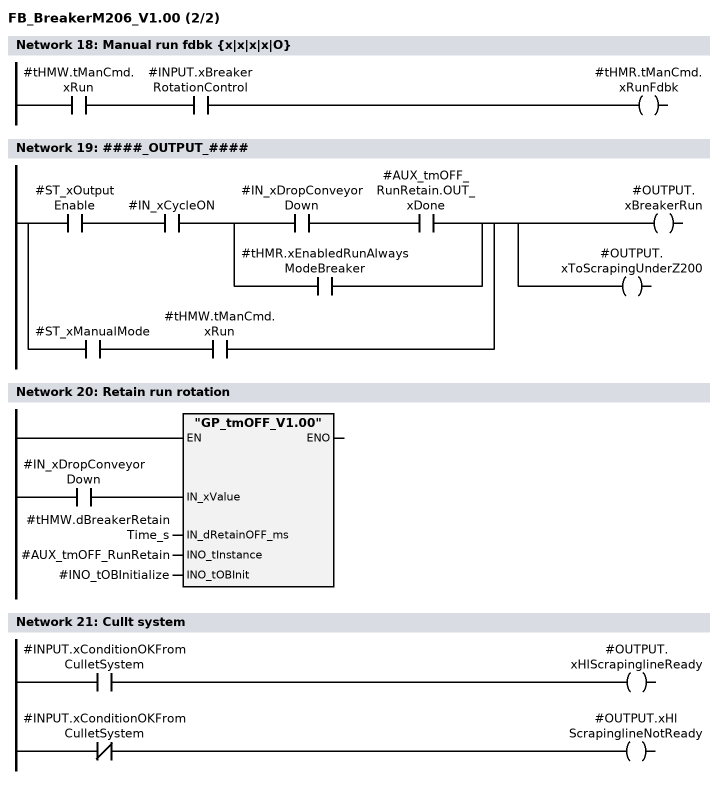
   RUNG wire#powerrail
      Contact( #tHMW.tManCmd.xRun )
      Contact( #INPUT.xBreakerRotationControl )
      Coil( #tHMR.tManCmd.xRunFdbk )
   END_RUNG
   // the same network as SCL:
   #tHMR.tManCmd.xRunFdbk := #tHMW.tManCmd.xRun AND #INPUT.xBreakerRotationControl;
END_REGION

REGION Network 19: ####_OUTPUT_####
   RUNG wire#powerrail
      Contact( #ST_xOutputEnable )
      Contact( #IN_xCycleON )
      wire#w1
      Contact( #IN_xDropConveyorDown )
      Contact( #AUX_tmOFF_RunRetain.OUT_xDone )
      wire#w2
      Coil( #OUTPUT.xBreakerRun )
   END_RUNG
   RUNG wire#w1
      Contact( #tHMR.xEnabledRunAlwaysModeBreaker )
   END_RUNG wire#w2
   RUNG wire#powerrail
      Contact( #ST_xManualMode )
      Contact( #tHMW.tManCmd.xRun )
   END_RUNG wire#w2
   RUNG wire#w2
      Coil( #OUTPUT.xToScrapingUnderZ200 )
   END_RUNG
   // the same network as SCL:
   #OUTPUT.xBreakerRun := (#ST_xOutputEnable AND #IN_xCycleON AND ((#IN_xDropConveyorDown AND #AUX_tmOFF_RunRetain.OUT_xDone) OR #tHMR.xEnabledRunAlwaysModeBreaker)) OR (#ST_xManualMode AND #tHMW.tManCmd.xRun);
   #OUTPUT.xToScrapingUnderZ200 := #OUTPUT.xBreakerRun;
END_REGION

REGION Network 20: Retain run rotation
   RUNG wire#powerrail
      "GP_tmOFF_V1.00"(IN_xValue := wire#w1, IN_dRetainOFF_ms := #tHMW.dBreakerRetainTime_s, INO_tInstance := #AUX_tmOFF_RunRetain, INO_tOBInit := #INO_tOBInitialize)
   END_RUNG
   RUNG wire#powerrail
      Contact( #IN_xDropConveyorDown )
   END_RUNG wire#w1
   // the same network as SCL:
   "GP_tmOFF_V1.00"(IN_xValue := #IN_xDropConveyorDown,
                    IN_dRetainOFF_ms := #tHMW.dBreakerRetainTime_s,
                    INO_tInstance := #AUX_tmOFF_RunRetain,
                    INO_tOBInit := #INO_tOBInitialize);
END_REGION

REGION Network 21: Cullt system
   RUNG wire#powerrail
      Contact( #INPUT.xConditionOKFromCulletSystem )
      Coil( #OUTPUT.xHlScrapinglineReady )
   END_RUNG
   RUNG wire#powerrail
      I_Contact( #INPUT.xConditionOKFromCulletSystem )
      Coil( #OUTPUT.xHlScrapinglineNotReady )
   END_RUNG
   // the same network as SCL:
   #OUTPUT.xHlScrapinglineReady := #INPUT.xConditionOKFromCulletSystem;
   #OUTPUT.xHlScrapinglineNotReady := NOT #INPUT.xConditionOKFromCulletSystem;
END_REGION
END_FUNCTION_BLOCK

// folder: 03_Programs_Logics/MCC1201/26_RollsConveyorZ200

FUNCTION_BLOCK "FB_Z200Conveyor_SinamicsMotor"   // FB26, LAD
{ S7_Optimized_Access := 'TRUE' }